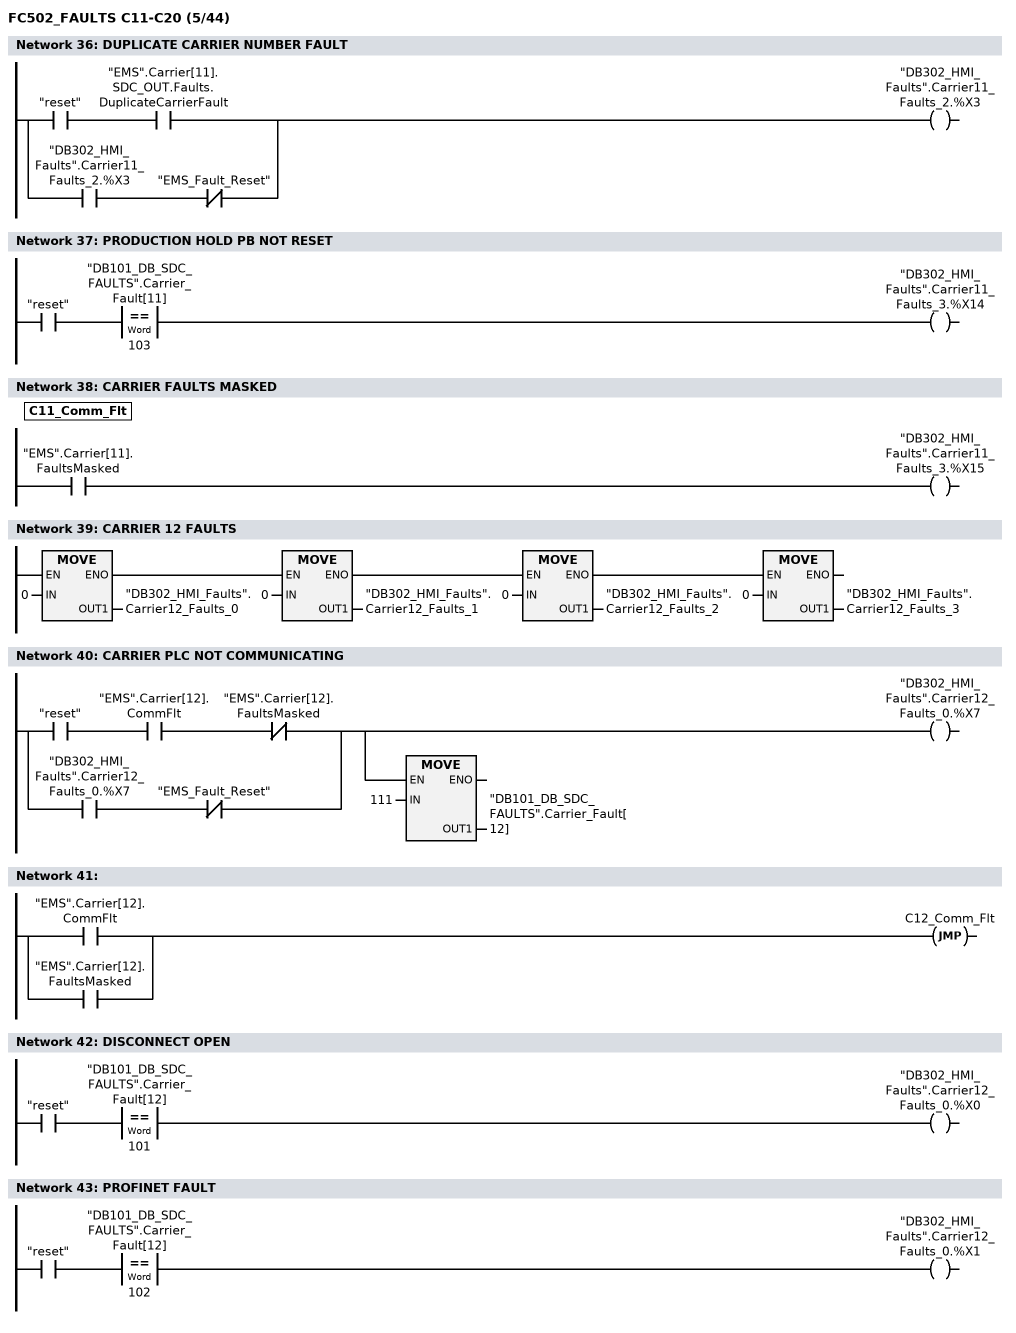
   RUNG wire#powerrail
      Contact( "reset" )
      Contact( "EMS".Carrier[11].SDC_OUT.Faults.DuplicateCarrierFault )
      wire#w1
      Coil( "DB302_HMI_Faults".Carrier11_Faults_2.%X3 )
   END_RUNG
   RUNG wire#powerrail
      Contact( "DB302_HMI_Faults".Carrier11_Faults_2.%X3 )
      I_Contact( "EMS_Fault_Reset" )
   END_RUNG wire#w1
   // the same network as SCL:
   "DB302_HMI_Faults".Carrier11_Faults_2.%X3 := ("reset" AND "EMS".Carrier[11].SDC_OUT.Faults.DuplicateCarrierFault) OR ("DB302_HMI_Faults".Carrier11_Faults_2.%X3 AND NOT "EMS_Fault_Reset");
END_REGION

REGION Network 37: PRODUCTION HOLD PB NOT RESET
   RUNG wire#powerrail
      Contact( "reset" )
      { S7_Templates := "SrcType := Word" } EQ_Contact(in1 := "DB101_DB_SDC_FAULTS".Carrier_Fault[11], in2 := 103)
      Coil( "DB302_HMI_Faults".Carrier11_Faults_3.%X14 )
   END_RUNG
   // the same network as SCL:
   "DB302_HMI_Faults".Carrier11_Faults_3.%X14 := "reset" AND ("DB101_DB_SDC_FAULTS".Carrier_Fault[11] = 103);
END_REGION

REGION Network 38: CARRIER FAULTS MASKED
   Label( C11_Comm_Flt )
   RUNG wire#powerrail
      Contact( "EMS".Carrier[11].FaultsMasked )
      Coil( "DB302_HMI_Faults".Carrier11_Faults_3.%X15 )
   END_RUNG
   // the same network as SCL:
   C11_Comm_Flt:
   "DB302_HMI_Faults".Carrier11_Faults_3.%X15 := "EMS".Carrier[11].FaultsMasked;
END_REGION

REGION Network 39: CARRIER 12 FAULTS
   RUNG wire#powerrail
      Move(in := 0, out1 => "DB302_HMI_Faults".Carrier12_Faults_0)
      Move(in := 0, out1 => "DB302_HMI_Faults".Carrier12_Faults_1)
      Move(in := 0, out1 => "DB302_HMI_Faults".Carrier12_Faults_2)
      Move(in := 0, out1 => "DB302_HMI_Faults".Carrier12_Faults_3)
   END_RUNG
   // the same network as SCL:
   "DB302_HMI_Faults".Carrier12_Faults_0 := 0;
   "DB302_HMI_Faults".Carrier12_Faults_1 := 0;
   "DB302_HMI_Faults".Carrier12_Faults_2 := 0;
   "DB302_HMI_Faults".Carrier12_Faults_3 := 0;
END_REGION

REGION Network 40: CARRIER PLC NOT COMMUNICATING
   RUNG wire#powerrail
      Contact( "reset" )
      Contact( "EMS".Carrier[12].CommFlt )
      I_Contact( "EMS".Carrier[12].FaultsMasked )
      wire#w1
      Coil( "DB302_HMI_Faults".Carrier12_Faults_0.%X7 )
   END_RUNG
   RUNG wire#powerrail
      Contact( "DB302_HMI_Faults".Carrier12_Faults_0.%X7 )
      I_Contact( "EMS_Fault_Reset" )
   END_RUNG wire#w1
   RUNG wire#w1
      Move(in := 111, out1 => "DB101_DB_SDC_FAULTS".Carrier_Fault[12])
   END_RUNG
   // the same network as SCL:
   "DB302_HMI_Faults".Carrier12_Faults_0.%X7 := ("reset" AND "EMS".Carrier[12].CommFlt AND NOT "EMS".Carrier[12].FaultsMasked) OR ("DB302_HMI_Faults".Carrier12_Faults_0.%X7 AND NOT "EMS_Fault_Reset");
   IF "DB302_HMI_Faults".Carrier12_Faults_0.%X7 THEN "DB101_DB_SDC_FAULTS".Carrier_Fault[12] := 111; END_IF;
END_REGION

REGION Network 41
   RUNG wire#powerrail
      Contact( "EMS".Carrier[12].CommFlt )
      wire#w1
      JumpCoil( C12_Comm_Flt )
   END_RUNG
   RUNG wire#powerrail
      Contact( "EMS".Carrier[12].FaultsMasked )
   END_RUNG wire#w1
   // the same network as SCL:
   IF "EMS".Carrier[12].CommFlt OR "EMS".Carrier[12].FaultsMasked THEN GOTO C12_Comm_Flt; END_IF;
END_REGION

REGION Network 42: DISCONNECT OPEN
   RUNG wire#powerrail
      Contact( "reset" )
      { S7_Templates := "SrcType := Word" } EQ_Contact(in1 := "DB101_DB_SDC_FAULTS".Carrier_Fault[12], in2 := 101)
      Coil( "DB302_HMI_Faults".Carrier12_Faults_0.%X0 )
   END_RUNG
   // the same network as SCL:
   "DB302_HMI_Faults".Carrier12_Faults_0.%X0 := "reset" AND ("DB101_DB_SDC_FAULTS".Carrier_Fault[12] = 101);
END_REGION

REGION Network 43: PROFINET FAULT
   RUNG wire#powerrail
      Contact( "reset" )
      { S7_Templates := "SrcType := Word" } EQ_Contact(in1 := "DB101_DB_SDC_FAULTS".Carrier_Fault[12], in2 := 102)
      Coil( "DB302_HMI_Faults".Carrier12_Faults_0.%X1 )
   END_RUNG
   // the same network as SCL:
   "DB302_HMI_Faults".Carrier12_Faults_0.%X1 := "reset" AND ("DB101_DB_SDC_FAULTS".Carrier_Fault[12] = 102);
END_REGION

REGION Network 44: CB2122 TRIPPED
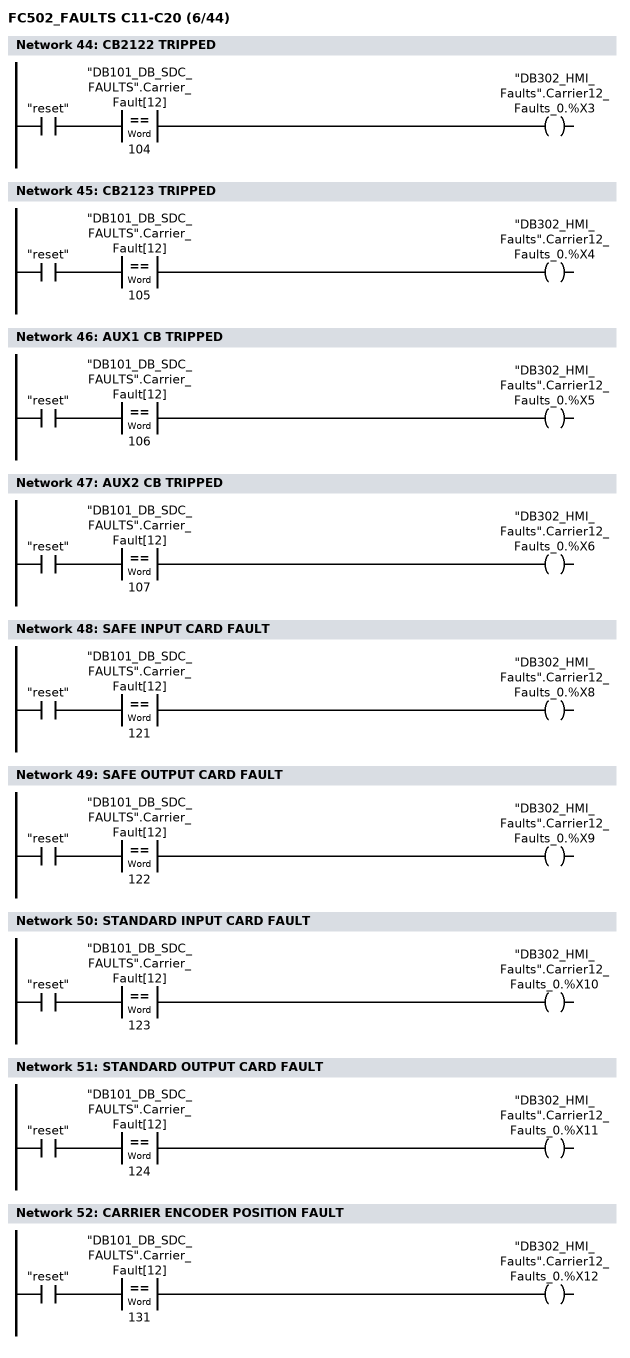
   RUNG wire#powerrail
      Contact( "reset" )
      { S7_Templates := "SrcType := Word" } EQ_Contact(in1 := "DB101_DB_SDC_FAULTS".Carrier_Fault[12], in2 := 104)
      Coil( "DB302_HMI_Faults".Carrier12_Faults_0.%X3 )
   END_RUNG
   // the same network as SCL:
   "DB302_HMI_Faults".Carrier12_Faults_0.%X3 := "reset" AND ("DB101_DB_SDC_FAULTS".Carrier_Fault[12] = 104);
END_REGION

REGION Network 45: CB2123 TRIPPED
   RUNG wire#powerrail
      Contact( "reset" )
      { S7_Templates := "SrcType := Word" } EQ_Contact(in1 := "DB101_DB_SDC_FAULTS".Carrier_Fault[12], in2 := 105)
      Coil( "DB302_HMI_Faults".Carrier12_Faults_0.%X4 )
   END_RUNG
   // the same network as SCL:
   "DB302_HMI_Faults".Carrier12_Faults_0.%X4 := "reset" AND ("DB101_DB_SDC_FAULTS".Carrier_Fault[12] = 105);
END_REGION

REGION Network 46: AUX1 CB TRIPPED
   RUNG wire#powerrail
      Contact( "reset" )
      { S7_Templates := "SrcType := Word" } EQ_Contact(in1 := "DB101_DB_SDC_FAULTS".Carrier_Fault[12], in2 := 106)
      Coil( "DB302_HMI_Faults".Carrier12_Faults_0.%X5 )
   END_RUNG
   // the same network as SCL:
   "DB302_HMI_Faults".Carrier12_Faults_0.%X5 := "reset" AND ("DB101_DB_SDC_FAULTS".Carrier_Fault[12] = 106);
END_REGION

REGION Network 47: AUX2 CB TRIPPED
   RUNG wire#powerrail
      Contact( "reset" )
      { S7_Templates := "SrcType := Word" } EQ_Contact(in1 := "DB101_DB_SDC_FAULTS".Carrier_Fault[12], in2 := 107)
      Coil( "DB302_HMI_Faults".Carrier12_Faults_0.%X6 )
   END_RUNG
   // the same network as SCL:
   "DB302_HMI_Faults".Carrier12_Faults_0.%X6 := "reset" AND ("DB101_DB_SDC_FAULTS".Carrier_Fault[12] = 107);
END_REGION

REGION Network 48: SAFE INPUT CARD FAULT
   RUNG wire#powerrail
      Contact( "reset" )
      { S7_Templates := "SrcType := Word" } EQ_Contact(in1 := "DB101_DB_SDC_FAULTS".Carrier_Fault[12], in2 := 121)
      Coil( "DB302_HMI_Faults".Carrier12_Faults_0.%X8 )
   END_RUNG
   // the same network as SCL:
   "DB302_HMI_Faults".Carrier12_Faults_0.%X8 := "reset" AND ("DB101_DB_SDC_FAULTS".Carrier_Fault[12] = 121);
END_REGION

REGION Network 49: SAFE OUTPUT CARD FAULT
   RUNG wire#powerrail
      Contact( "reset" )
      { S7_Templates := "SrcType := Word" } EQ_Contact(in1 := "DB101_DB_SDC_FAULTS".Carrier_Fault[12], in2 := 122)
      Coil( "DB302_HMI_Faults".Carrier12_Faults_0.%X9 )
   END_RUNG
   // the same network as SCL:
   "DB302_HMI_Faults".Carrier12_Faults_0.%X9 := "reset" AND ("DB101_DB_SDC_FAULTS".Carrier_Fault[12] = 122);
END_REGION

REGION Network 50: STANDARD INPUT CARD FAULT
   RUNG wire#powerrail
      Contact( "reset" )
      { S7_Templates := "SrcType := Word" } EQ_Contact(in1 := "DB101_DB_SDC_FAULTS".Carrier_Fault[12], in2 := 123)
      Coil( "DB302_HMI_Faults".Carrier12_Faults_0.%X10 )
   END_RUNG
   // the same network as SCL:
   "DB302_HMI_Faults".Carrier12_Faults_0.%X10 := "reset" AND ("DB101_DB_SDC_FAULTS".Carrier_Fault[12] = 123);
END_REGION

REGION Network 51: STANDARD OUTPUT CARD FAULT
   RUNG wire#powerrail
      Contact( "reset" )
      { S7_Templates := "SrcType := Word" } EQ_Contact(in1 := "DB101_DB_SDC_FAULTS".Carrier_Fault[12], in2 := 124)
      Coil( "DB302_HMI_Faults".Carrier12_Faults_0.%X11 )
   END_RUNG
   // the same network as SCL:
   "DB302_HMI_Faults".Carrier12_Faults_0.%X11 := "reset" AND ("DB101_DB_SDC_FAULTS".Carrier_Fault[12] = 124);
END_REGION

REGION Network 52: CARRIER ENCODER POSITION FAULT
   RUNG wire#powerrail
      Contact( "reset" )
      { S7_Templates := "SrcType := Word" } EQ_Contact(in1 := "DB101_DB_SDC_FAULTS".Carrier_Fault[12], in2 := 131)
      Coil( "DB302_HMI_Faults".Carrier12_Faults_0.%X12 )
   END_RUNG
   // the same network as SCL:
   "DB302_HMI_Faults".Carrier12_Faults_0.%X12 := "reset" AND ("DB101_DB_SDC_FAULTS".Carrier_Fault[12] = 131);
END_REGION

REGION Network 53: CARRIER ENCODER INTERNAL ERROR
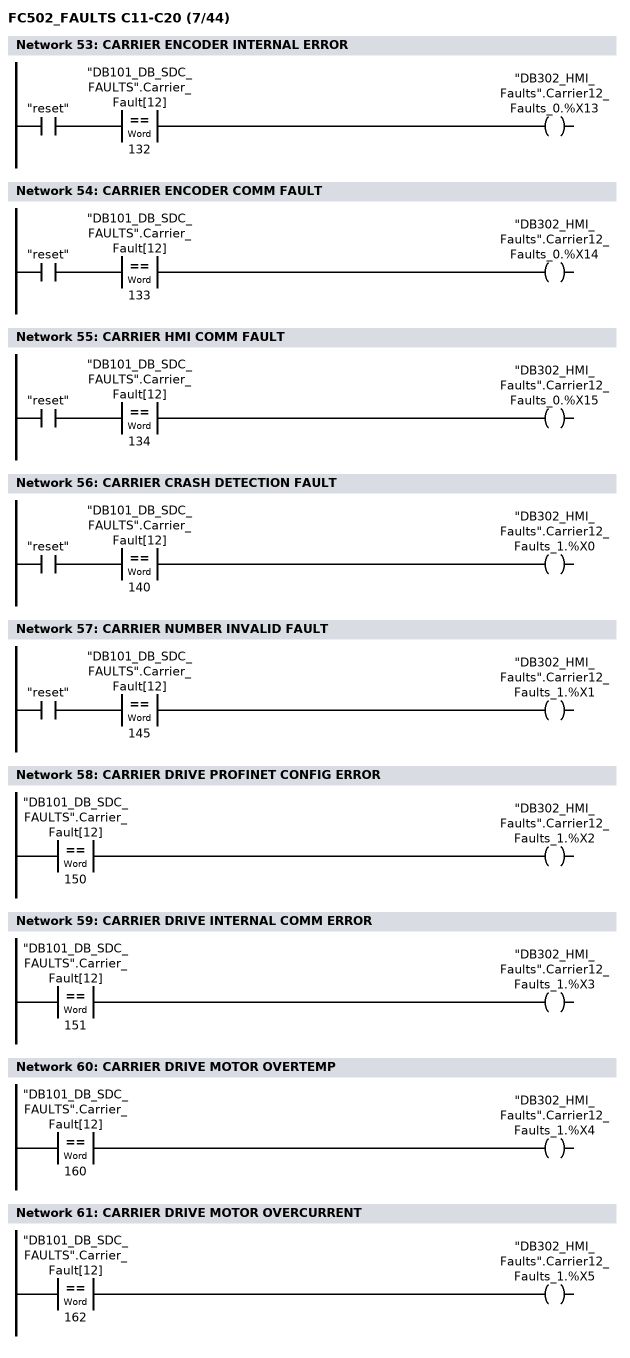
   RUNG wire#powerrail
      Contact( "reset" )
      { S7_Templates := "SrcType := Word" } EQ_Contact(in1 := "DB101_DB_SDC_FAULTS".Carrier_Fault[12], in2 := 132)
      Coil( "DB302_HMI_Faults".Carrier12_Faults_0.%X13 )
   END_RUNG
   // the same network as SCL:
   "DB302_HMI_Faults".Carrier12_Faults_0.%X13 := "reset" AND ("DB101_DB_SDC_FAULTS".Carrier_Fault[12] = 132);
END_REGION

REGION Network 54: CARRIER ENCODER COMM FAULT
   RUNG wire#powerrail
      Contact( "reset" )
      { S7_Templates := "SrcType := Word" } EQ_Contact(in1 := "DB101_DB_SDC_FAULTS".Carrier_Fault[12], in2 := 133)
      Coil( "DB302_HMI_Faults".Carrier12_Faults_0.%X14 )
   END_RUNG
   // the same network as SCL:
   "DB302_HMI_Faults".Carrier12_Faults_0.%X14 := "reset" AND ("DB101_DB_SDC_FAULTS".Carrier_Fault[12] = 133);
END_REGION

REGION Network 55: CARRIER HMI COMM FAULT
   RUNG wire#powerrail
      Contact( "reset" )
      { S7_Templates := "SrcType := Word" } EQ_Contact(in1 := "DB101_DB_SDC_FAULTS".Carrier_Fault[12], in2 := 134)
      Coil( "DB302_HMI_Faults".Carrier12_Faults_0.%X15 )
   END_RUNG
   // the same network as SCL:
   "DB302_HMI_Faults".Carrier12_Faults_0.%X15 := "reset" AND ("DB101_DB_SDC_FAULTS".Carrier_Fault[12] = 134);
END_REGION

REGION Network 56: CARRIER CRASH DETECTION FAULT
   RUNG wire#powerrail
      Contact( "reset" )
      { S7_Templates := "SrcType := Word" } EQ_Contact(in1 := "DB101_DB_SDC_FAULTS".Carrier_Fault[12], in2 := 140)
      Coil( "DB302_HMI_Faults".Carrier12_Faults_1.%X0 )
   END_RUNG
   // the same network as SCL:
   "DB302_HMI_Faults".Carrier12_Faults_1.%X0 := "reset" AND ("DB101_DB_SDC_FAULTS".Carrier_Fault[12] = 140);
END_REGION

REGION Network 57: CARRIER NUMBER INVALID FAULT
   RUNG wire#powerrail
      Contact( "reset" )
      { S7_Templates := "SrcType := Word" } EQ_Contact(in1 := "DB101_DB_SDC_FAULTS".Carrier_Fault[12], in2 := 145)
      Coil( "DB302_HMI_Faults".Carrier12_Faults_1.%X1 )
   END_RUNG
   // the same network as SCL:
   "DB302_HMI_Faults".Carrier12_Faults_1.%X1 := "reset" AND ("DB101_DB_SDC_FAULTS".Carrier_Fault[12] = 145);
END_REGION

REGION Network 58: CARRIER DRIVE PROFINET CONFIG ERROR
   RUNG wire#powerrail
      { S7_Templates := "SrcType := Word" } EQ_Contact(in1 := "DB101_DB_SDC_FAULTS".Carrier_Fault[12], in2 := 150)
      Coil( "DB302_HMI_Faults".Carrier12_Faults_1.%X2 )
   END_RUNG
   // the same network as SCL:
   "DB302_HMI_Faults".Carrier12_Faults_1.%X2 := "DB101_DB_SDC_FAULTS".Carrier_Fault[12] = 150;
END_REGION

REGION Network 59: CARRIER DRIVE INTERNAL COMM ERROR
   RUNG wire#powerrail
      { S7_Templates := "SrcType := Word" } EQ_Contact(in1 := "DB101_DB_SDC_FAULTS".Carrier_Fault[12], in2 := 151)
      Coil( "DB302_HMI_Faults".Carrier12_Faults_1.%X3 )
   END_RUNG
   // the same network as SCL:
   "DB302_HMI_Faults".Carrier12_Faults_1.%X3 := "DB101_DB_SDC_FAULTS".Carrier_Fault[12] = 151;
END_REGION

REGION Network 60: CARRIER DRIVE MOTOR OVERTEMP
   RUNG wire#powerrail
      { S7_Templates := "SrcType := Word" } EQ_Contact(in1 := "DB101_DB_SDC_FAULTS".Carrier_Fault[12], in2 := 160)
      Coil( "DB302_HMI_Faults".Carrier12_Faults_1.%X4 )
   END_RUNG
   // the same network as SCL:
   "DB302_HMI_Faults".Carrier12_Faults_1.%X4 := "DB101_DB_SDC_FAULTS".Carrier_Fault[12] = 160;
END_REGION

REGION Network 61: CARRIER DRIVE MOTOR OVERCURRENT
   RUNG wire#powerrail
      { S7_Templates := "SrcType := Word" } EQ_Contact(in1 := "DB101_DB_SDC_FAULTS".Carrier_Fault[12], in2 := 162)
      Coil( "DB302_HMI_Faults".Carrier12_Faults_1.%X5 )
   END_RUNG
   // the same network as SCL:
   "DB302_HMI_Faults".Carrier12_Faults_1.%X5 := "DB101_DB_SDC_FAULTS".Carrier_Fault[12] = 162;
END_REGION

REGION Network 62: CARRIER DRIVE INFEED OR POWER UNIT NOT READY
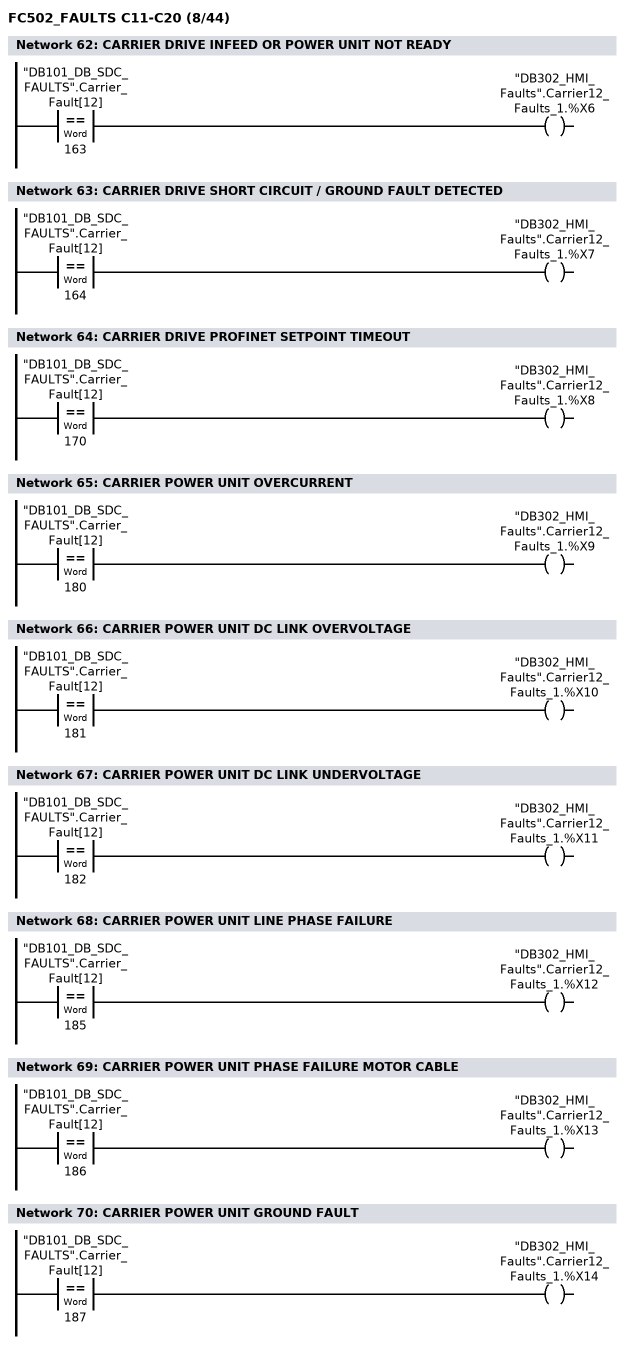
   RUNG wire#powerrail
      { S7_Templates := "SrcType := Word" } EQ_Contact(in1 := "DB101_DB_SDC_FAULTS".Carrier_Fault[12], in2 := 163)
      Coil( "DB302_HMI_Faults".Carrier12_Faults_1.%X6 )
   END_RUNG
   // the same network as SCL:
   "DB302_HMI_Faults".Carrier12_Faults_1.%X6 := "DB101_DB_SDC_FAULTS".Carrier_Fault[12] = 163;
END_REGION

REGION Network 63: CARRIER DRIVE SHORT CIRCUIT / GROUND FAULT DETECTED
   RUNG wire#powerrail
      { S7_Templates := "SrcType := Word" } EQ_Contact(in1 := "DB101_DB_SDC_FAULTS".Carrier_Fault[12], in2 := 164)
      Coil( "DB302_HMI_Faults".Carrier12_Faults_1.%X7 )
   END_RUNG
   // the same network as SCL:
   "DB302_HMI_Faults".Carrier12_Faults_1.%X7 := "DB101_DB_SDC_FAULTS".Carrier_Fault[12] = 164;
END_REGION

REGION Network 64: CARRIER DRIVE PROFINET SETPOINT TIMEOUT
   RUNG wire#powerrail
      { S7_Templates := "SrcType := Word" } EQ_Contact(in1 := "DB101_DB_SDC_FAULTS".Carrier_Fault[12], in2 := 170)
      Coil( "DB302_HMI_Faults".Carrier12_Faults_1.%X8 )
   END_RUNG
   // the same network as SCL:
   "DB302_HMI_Faults".Carrier12_Faults_1.%X8 := "DB101_DB_SDC_FAULTS".Carrier_Fault[12] = 170;
END_REGION

REGION Network 65: CARRIER POWER UNIT OVERCURRENT
   RUNG wire#powerrail
      { S7_Templates := "SrcType := Word" } EQ_Contact(in1 := "DB101_DB_SDC_FAULTS".Carrier_Fault[12], in2 := 180)
      Coil( "DB302_HMI_Faults".Carrier12_Faults_1.%X9 )
   END_RUNG
   // the same network as SCL:
   "DB302_HMI_Faults".Carrier12_Faults_1.%X9 := "DB101_DB_SDC_FAULTS".Carrier_Fault[12] = 180;
END_REGION

REGION Network 66: CARRIER POWER UNIT DC LINK OVERVOLTAGE
   RUNG wire#powerrail
      { S7_Templates := "SrcType := Word" } EQ_Contact(in1 := "DB101_DB_SDC_FAULTS".Carrier_Fault[12], in2 := 181)
      Coil( "DB302_HMI_Faults".Carrier12_Faults_1.%X10 )
   END_RUNG
   // the same network as SCL:
   "DB302_HMI_Faults".Carrier12_Faults_1.%X10 := "DB101_DB_SDC_FAULTS".Carrier_Fault[12] = 181;
END_REGION

REGION Network 67: CARRIER POWER UNIT DC LINK UNDERVOLTAGE
   RUNG wire#powerrail
      { S7_Templates := "SrcType := Word" } EQ_Contact(in1 := "DB101_DB_SDC_FAULTS".Carrier_Fault[12], in2 := 182)
      Coil( "DB302_HMI_Faults".Carrier12_Faults_1.%X11 )
   END_RUNG
   // the same network as SCL:
   "DB302_HMI_Faults".Carrier12_Faults_1.%X11 := "DB101_DB_SDC_FAULTS".Carrier_Fault[12] = 182;
END_REGION

REGION Network 68: CARRIER POWER UNIT LINE PHASE FAILURE
   RUNG wire#powerrail
      { S7_Templates := "SrcType := Word" } EQ_Contact(in1 := "DB101_DB_SDC_FAULTS".Carrier_Fault[12], in2 := 185)
      Coil( "DB302_HMI_Faults".Carrier12_Faults_1.%X12 )
   END_RUNG
   // the same network as SCL:
   "DB302_HMI_Faults".Carrier12_Faults_1.%X12 := "DB101_DB_SDC_FAULTS".Carrier_Fault[12] = 185;
END_REGION

REGION Network 69: CARRIER POWER UNIT PHASE FAILURE MOTOR CABLE
   RUNG wire#powerrail
      { S7_Templates := "SrcType := Word" } EQ_Contact(in1 := "DB101_DB_SDC_FAULTS".Carrier_Fault[12], in2 := 186)
      Coil( "DB302_HMI_Faults".Carrier12_Faults_1.%X13 )
   END_RUNG
   // the same network as SCL:
   "DB302_HMI_Faults".Carrier12_Faults_1.%X13 := "DB101_DB_SDC_FAULTS".Carrier_Fault[12] = 186;
END_REGION

REGION Network 70: CARRIER POWER UNIT GROUND FAULT
   RUNG wire#powerrail
      { S7_Templates := "SrcType := Word" } EQ_Contact(in1 := "DB101_DB_SDC_FAULTS".Carrier_Fault[12], in2 := 187)
      Coil( "DB302_HMI_Faults".Carrier12_Faults_1.%X14 )
   END_RUNG
   // the same network as SCL:
   "DB302_HMI_Faults".Carrier12_Faults_1.%X14 := "DB101_DB_SDC_FAULTS".Carrier_Fault[12] = 187;
END_REGION

REGION Network 71: CARRIER MOTION OFF FAULT
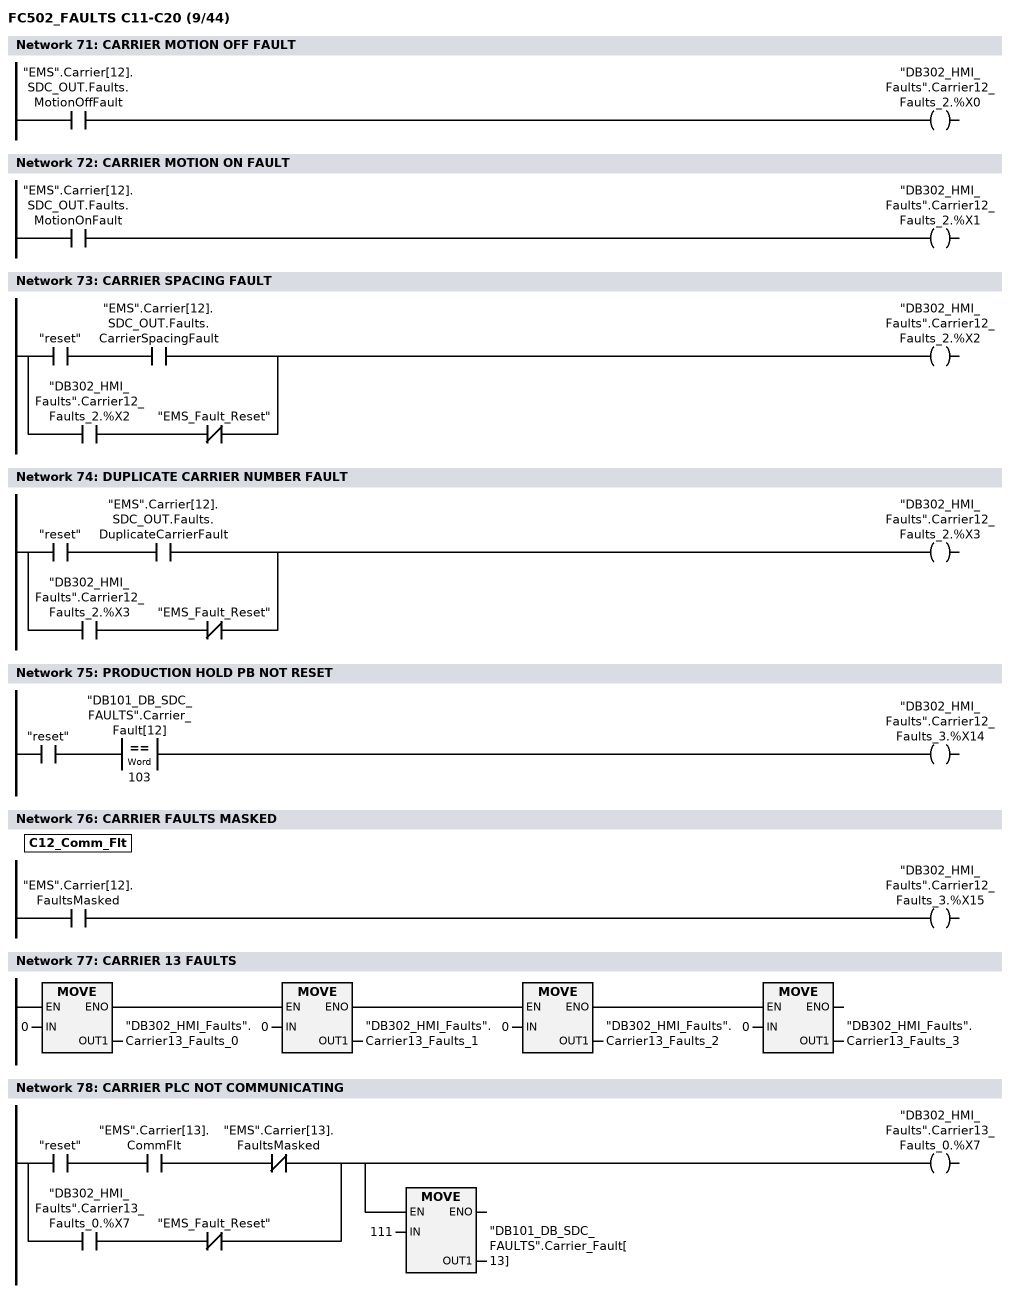
   RUNG wire#powerrail
      Contact( "EMS".Carrier[12].SDC_OUT.Faults.MotionOffFault )
      Coil( "DB302_HMI_Faults".Carrier12_Faults_2.%X0 )
   END_RUNG
   // the same network as SCL:
   "DB302_HMI_Faults".Carrier12_Faults_2.%X0 := "EMS".Carrier[12].SDC_OUT.Faults.MotionOffFault;
END_REGION

REGION Network 72: CARRIER MOTION ON FAULT
   RUNG wire#powerrail
      Contact( "EMS".Carrier[12].SDC_OUT.Faults.MotionOnFault )
      Coil( "DB302_HMI_Faults".Carrier12_Faults_2.%X1 )
   END_RUNG
   // the same network as SCL:
   "DB302_HMI_Faults".Carrier12_Faults_2.%X1 := "EMS".Carrier[12].SDC_OUT.Faults.MotionOnFault;
END_REGION

REGION Network 73: CARRIER SPACING FAULT
   RUNG wire#powerrail
      Contact( "reset" )
      Contact( "EMS".Carrier[12].SDC_OUT.Faults.CarrierSpacingFault )
      wire#w1
      Coil( "DB302_HMI_Faults".Carrier12_Faults_2.%X2 )
   END_RUNG
   RUNG wire#powerrail
      Contact( "DB302_HMI_Faults".Carrier12_Faults_2.%X2 )
      I_Contact( "EMS_Fault_Reset" )
   END_RUNG wire#w1
   // the same network as SCL:
   "DB302_HMI_Faults".Carrier12_Faults_2.%X2 := ("reset" AND "EMS".Carrier[12].SDC_OUT.Faults.CarrierSpacingFault) OR ("DB302_HMI_Faults".Carrier12_Faults_2.%X2 AND NOT "EMS_Fault_Reset");
END_REGION

REGION Network 74: DUPLICATE CARRIER NUMBER FAULT
   RUNG wire#powerrail
      Contact( "reset" )
      Contact( "EMS".Carrier[12].SDC_OUT.Faults.DuplicateCarrierFault )
      wire#w1
      Coil( "DB302_HMI_Faults".Carrier12_Faults_2.%X3 )
   END_RUNG
   RUNG wire#powerrail
      Contact( "DB302_HMI_Faults".Carrier12_Faults_2.%X3 )
      I_Contact( "EMS_Fault_Reset" )
   END_RUNG wire#w1
   // the same network as SCL:
   "DB302_HMI_Faults".Carrier12_Faults_2.%X3 := ("reset" AND "EMS".Carrier[12].SDC_OUT.Faults.DuplicateCarrierFault) OR ("DB302_HMI_Faults".Carrier12_Faults_2.%X3 AND NOT "EMS_Fault_Reset");
END_REGION

REGION Network 75: PRODUCTION HOLD PB NOT RESET
   RUNG wire#powerrail
      Contact( "reset" )
      { S7_Templates := "SrcType := Word" } EQ_Contact(in1 := "DB101_DB_SDC_FAULTS".Carrier_Fault[12], in2 := 103)
      Coil( "DB302_HMI_Faults".Carrier12_Faults_3.%X14 )
   END_RUNG
   // the same network as SCL:
   "DB302_HMI_Faults".Carrier12_Faults_3.%X14 := "reset" AND ("DB101_DB_SDC_FAULTS".Carrier_Fault[12] = 103);
END_REGION

REGION Network 76: CARRIER FAULTS MASKED
   Label( C12_Comm_Flt )
   RUNG wire#powerrail
      Contact( "EMS".Carrier[12].FaultsMasked )
      Coil( "DB302_HMI_Faults".Carrier12_Faults_3.%X15 )
   END_RUNG
   // the same network as SCL:
   C12_Comm_Flt:
   "DB302_HMI_Faults".Carrier12_Faults_3.%X15 := "EMS".Carrier[12].FaultsMasked;
END_REGION

REGION Network 77: CARRIER 13 FAULTS
   RUNG wire#powerrail
      Move(in := 0, out1 => "DB302_HMI_Faults".Carrier13_Faults_0)
      Move(in := 0, out1 => "DB302_HMI_Faults".Carrier13_Faults_1)
      Move(in := 0, out1 => "DB302_HMI_Faults".Carrier13_Faults_2)
      Move(in := 0, out1 => "DB302_HMI_Faults".Carrier13_Faults_3)
   END_RUNG
   // the same network as SCL:
   "DB302_HMI_Faults".Carrier13_Faults_0 := 0;
   "DB302_HMI_Faults".Carrier13_Faults_1 := 0;
   "DB302_HMI_Faults".Carrier13_Faults_2 := 0;
   "DB302_HMI_Faults".Carrier13_Faults_3 := 0;
END_REGION

REGION Network 78: CARRIER PLC NOT COMMUNICATING
   RUNG wire#powerrail
      Contact( "reset" )
      Contact( "EMS".Carrier[13].CommFlt )
      I_Contact( "EMS".Carrier[13].FaultsMasked )
      wire#w1
      Coil( "DB302_HMI_Faults".Carrier13_Faults_0.%X7 )
   END_RUNG
   RUNG wire#powerrail
      Contact( "DB302_HMI_Faults".Carrier13_Faults_0.%X7 )
      I_Contact( "EMS_Fault_Reset" )
   END_RUNG wire#w1
   RUNG wire#w1
      Move(in := 111, out1 => "DB101_DB_SDC_FAULTS".Carrier_Fault[13])
   END_RUNG
   // the same network as SCL:
   "DB302_HMI_Faults".Carrier13_Faults_0.%X7 := ("reset" AND "EMS".Carrier[13].CommFlt AND NOT "EMS".Carrier[13].FaultsMasked) OR ("DB302_HMI_Faults".Carrier13_Faults_0.%X7 AND NOT "EMS_Fault_Reset");
   IF "DB302_HMI_Faults".Carrier13_Faults_0.%X7 THEN "DB101_DB_SDC_FAULTS".Carrier_Fault[13] := 111; END_IF;
END_REGION

REGION Network 79
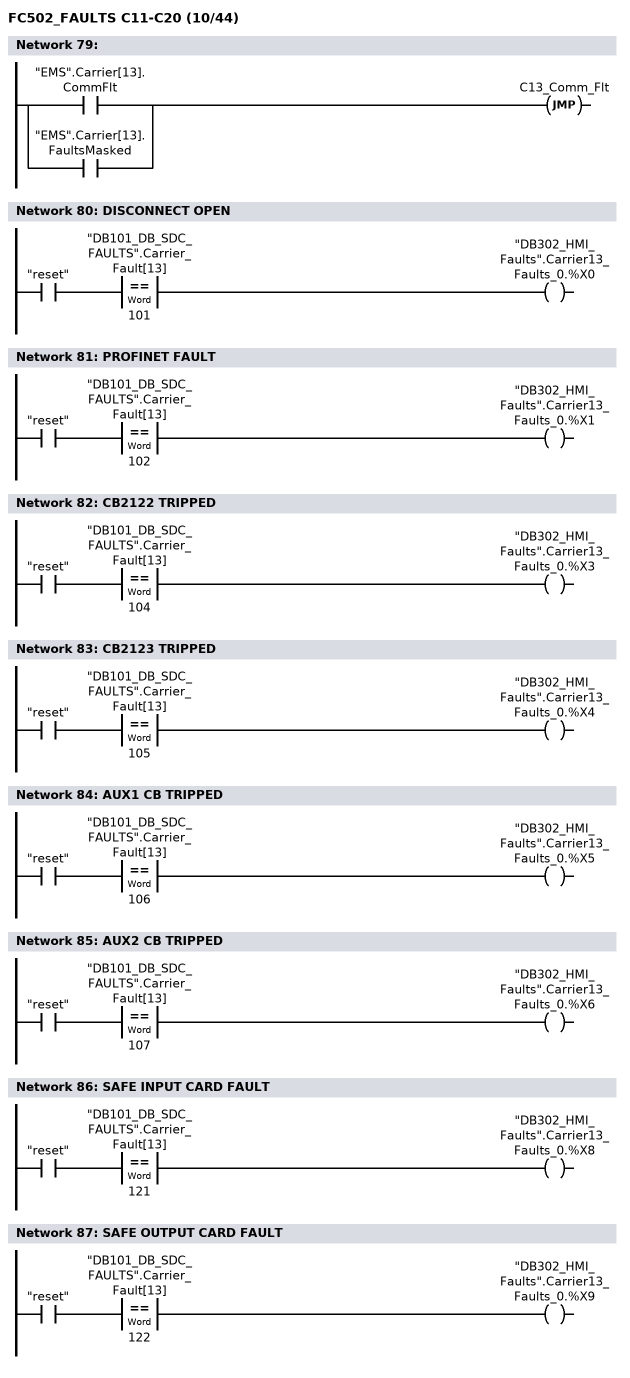
   RUNG wire#powerrail
      Contact( "EMS".Carrier[13].CommFlt )
      wire#w1
      JumpCoil( C13_Comm_Flt )
   END_RUNG
   RUNG wire#powerrail
      Contact( "EMS".Carrier[13].FaultsMasked )
   END_RUNG wire#w1
   // the same network as SCL:
   IF "EMS".Carrier[13].CommFlt OR "EMS".Carrier[13].FaultsMasked THEN GOTO C13_Comm_Flt; END_IF;
END_REGION

REGION Network 80: DISCONNECT OPEN
   RUNG wire#powerrail
      Contact( "reset" )
      { S7_Templates := "SrcType := Word" } EQ_Contact(in1 := "DB101_DB_SDC_FAULTS".Carrier_Fault[13], in2 := 101)
      Coil( "DB302_HMI_Faults".Carrier13_Faults_0.%X0 )
   END_RUNG
   // the same network as SCL:
   "DB302_HMI_Faults".Carrier13_Faults_0.%X0 := "reset" AND ("DB101_DB_SDC_FAULTS".Carrier_Fault[13] = 101);
END_REGION

REGION Network 81: PROFINET FAULT
   RUNG wire#powerrail
      Contact( "reset" )
      { S7_Templates := "SrcType := Word" } EQ_Contact(in1 := "DB101_DB_SDC_FAULTS".Carrier_Fault[13], in2 := 102)
      Coil( "DB302_HMI_Faults".Carrier13_Faults_0.%X1 )
   END_RUNG
   // the same network as SCL:
   "DB302_HMI_Faults".Carrier13_Faults_0.%X1 := "reset" AND ("DB101_DB_SDC_FAULTS".Carrier_Fault[13] = 102);
END_REGION

REGION Network 82: CB2122 TRIPPED
   RUNG wire#powerrail
      Contact( "reset" )
      { S7_Templates := "SrcType := Word" } EQ_Contact(in1 := "DB101_DB_SDC_FAULTS".Carrier_Fault[13], in2 := 104)
      Coil( "DB302_HMI_Faults".Carrier13_Faults_0.%X3 )
   END_RUNG
   // the same network as SCL:
   "DB302_HMI_Faults".Carrier13_Faults_0.%X3 := "reset" AND ("DB101_DB_SDC_FAULTS".Carrier_Fault[13] = 104);
END_REGION

REGION Network 83: CB2123 TRIPPED
   RUNG wire#powerrail
      Contact( "reset" )
      { S7_Templates := "SrcType := Word" } EQ_Contact(in1 := "DB101_DB_SDC_FAULTS".Carrier_Fault[13], in2 := 105)
      Coil( "DB302_HMI_Faults".Carrier13_Faults_0.%X4 )
   END_RUNG
   // the same network as SCL:
   "DB302_HMI_Faults".Carrier13_Faults_0.%X4 := "reset" AND ("DB101_DB_SDC_FAULTS".Carrier_Fault[13] = 105);
END_REGION

REGION Network 84: AUX1 CB TRIPPED
   RUNG wire#powerrail
      Contact( "reset" )
      { S7_Templates := "SrcType := Word" } EQ_Contact(in1 := "DB101_DB_SDC_FAULTS".Carrier_Fault[13], in2 := 106)
      Coil( "DB302_HMI_Faults".Carrier13_Faults_0.%X5 )
   END_RUNG
   // the same network as SCL:
   "DB302_HMI_Faults".Carrier13_Faults_0.%X5 := "reset" AND ("DB101_DB_SDC_FAULTS".Carrier_Fault[13] = 106);
END_REGION

REGION Network 85: AUX2 CB TRIPPED
   RUNG wire#powerrail
      Contact( "reset" )
      { S7_Templates := "SrcType := Word" } EQ_Contact(in1 := "DB101_DB_SDC_FAULTS".Carrier_Fault[13], in2 := 107)
      Coil( "DB302_HMI_Faults".Carrier13_Faults_0.%X6 )
   END_RUNG
   // the same network as SCL:
   "DB302_HMI_Faults".Carrier13_Faults_0.%X6 := "reset" AND ("DB101_DB_SDC_FAULTS".Carrier_Fault[13] = 107);
END_REGION

REGION Network 86: SAFE INPUT CARD FAULT
   RUNG wire#powerrail
      Contact( "reset" )
      { S7_Templates := "SrcType := Word" } EQ_Contact(in1 := "DB101_DB_SDC_FAULTS".Carrier_Fault[13], in2 := 121)
      Coil( "DB302_HMI_Faults".Carrier13_Faults_0.%X8 )
   END_RUNG
   // the same network as SCL:
   "DB302_HMI_Faults".Carrier13_Faults_0.%X8 := "reset" AND ("DB101_DB_SDC_FAULTS".Carrier_Fault[13] = 121);
END_REGION

REGION Network 87: SAFE OUTPUT CARD FAULT
   RUNG wire#powerrail
      Contact( "reset" )
      { S7_Templates := "SrcType := Word" } EQ_Contact(in1 := "DB101_DB_SDC_FAULTS".Carrier_Fault[13], in2 := 122)
      Coil( "DB302_HMI_Faults".Carrier13_Faults_0.%X9 )
   END_RUNG
   // the same network as SCL:
   "DB302_HMI_Faults".Carrier13_Faults_0.%X9 := "reset" AND ("DB101_DB_SDC_FAULTS".Carrier_Fault[13] = 122);
END_REGION

REGION Network 88: STANDARD INPUT CARD FAULT
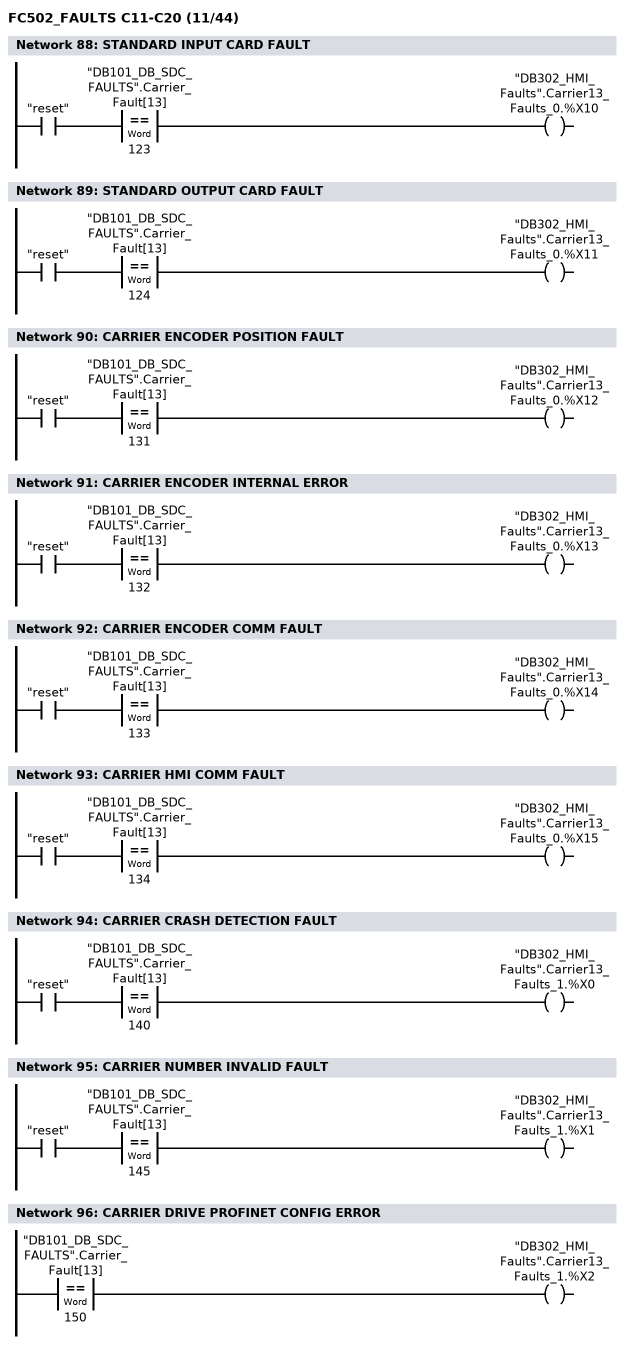
   RUNG wire#powerrail
      Contact( "reset" )
      { S7_Templates := "SrcType := Word" } EQ_Contact(in1 := "DB101_DB_SDC_FAULTS".Carrier_Fault[13], in2 := 123)
      Coil( "DB302_HMI_Faults".Carrier13_Faults_0.%X10 )
   END_RUNG
   // the same network as SCL:
   "DB302_HMI_Faults".Carrier13_Faults_0.%X10 := "reset" AND ("DB101_DB_SDC_FAULTS".Carrier_Fault[13] = 123);
END_REGION

REGION Network 89: STANDARD OUTPUT CARD FAULT
   RUNG wire#powerrail
      Contact( "reset" )
      { S7_Templates := "SrcType := Word" } EQ_Contact(in1 := "DB101_DB_SDC_FAULTS".Carrier_Fault[13], in2 := 124)
      Coil( "DB302_HMI_Faults".Carrier13_Faults_0.%X11 )
   END_RUNG
   // the same network as SCL:
   "DB302_HMI_Faults".Carrier13_Faults_0.%X11 := "reset" AND ("DB101_DB_SDC_FAULTS".Carrier_Fault[13] = 124);
END_REGION

REGION Network 90: CARRIER ENCODER POSITION FAULT
   RUNG wire#powerrail
      Contact( "reset" )
      { S7_Templates := "SrcType := Word" } EQ_Contact(in1 := "DB101_DB_SDC_FAULTS".Carrier_Fault[13], in2 := 131)
      Coil( "DB302_HMI_Faults".Carrier13_Faults_0.%X12 )
   END_RUNG
   // the same network as SCL:
   "DB302_HMI_Faults".Carrier13_Faults_0.%X12 := "reset" AND ("DB101_DB_SDC_FAULTS".Carrier_Fault[13] = 131);
END_REGION

REGION Network 91: CARRIER ENCODER INTERNAL ERROR
   RUNG wire#powerrail
      Contact( "reset" )
      { S7_Templates := "SrcType := Word" } EQ_Contact(in1 := "DB101_DB_SDC_FAULTS".Carrier_Fault[13], in2 := 132)
      Coil( "DB302_HMI_Faults".Carrier13_Faults_0.%X13 )
   END_RUNG
   // the same network as SCL:
   "DB302_HMI_Faults".Carrier13_Faults_0.%X13 := "reset" AND ("DB101_DB_SDC_FAULTS".Carrier_Fault[13] = 132);
END_REGION

REGION Network 92: CARRIER ENCODER COMM FAULT
   RUNG wire#powerrail
      Contact( "reset" )
      { S7_Templates := "SrcType := Word" } EQ_Contact(in1 := "DB101_DB_SDC_FAULTS".Carrier_Fault[13], in2 := 133)
      Coil( "DB302_HMI_Faults".Carrier13_Faults_0.%X14 )
   END_RUNG
   // the same network as SCL:
   "DB302_HMI_Faults".Carrier13_Faults_0.%X14 := "reset" AND ("DB101_DB_SDC_FAULTS".Carrier_Fault[13] = 133);
END_REGION

REGION Network 93: CARRIER HMI COMM FAULT
   RUNG wire#powerrail
      Contact( "reset" )
      { S7_Templates := "SrcType := Word" } EQ_Contact(in1 := "DB101_DB_SDC_FAULTS".Carrier_Fault[13], in2 := 134)
      Coil( "DB302_HMI_Faults".Carrier13_Faults_0.%X15 )
   END_RUNG
   // the same network as SCL:
   "DB302_HMI_Faults".Carrier13_Faults_0.%X15 := "reset" AND ("DB101_DB_SDC_FAULTS".Carrier_Fault[13] = 134);
END_REGION

REGION Network 94: CARRIER CRASH DETECTION FAULT
   RUNG wire#powerrail
      Contact( "reset" )
      { S7_Templates := "SrcType := Word" } EQ_Contact(in1 := "DB101_DB_SDC_FAULTS".Carrier_Fault[13], in2 := 140)
      Coil( "DB302_HMI_Faults".Carrier13_Faults_1.%X0 )
   END_RUNG
   // the same network as SCL:
   "DB302_HMI_Faults".Carrier13_Faults_1.%X0 := "reset" AND ("DB101_DB_SDC_FAULTS".Carrier_Fault[13] = 140);
END_REGION

REGION Network 95: CARRIER NUMBER INVALID FAULT
   RUNG wire#powerrail
      Contact( "reset" )
      { S7_Templates := "SrcType := Word" } EQ_Contact(in1 := "DB101_DB_SDC_FAULTS".Carrier_Fault[13], in2 := 145)
      Coil( "DB302_HMI_Faults".Carrier13_Faults_1.%X1 )
   END_RUNG
   // the same network as SCL:
   "DB302_HMI_Faults".Carrier13_Faults_1.%X1 := "reset" AND ("DB101_DB_SDC_FAULTS".Carrier_Fault[13] = 145);
END_REGION

REGION Network 96: CARRIER DRIVE PROFINET CONFIG ERROR
   RUNG wire#powerrail
      { S7_Templates := "SrcType := Word" } EQ_Contact(in1 := "DB101_DB_SDC_FAULTS".Carrier_Fault[13], in2 := 150)
      Coil( "DB302_HMI_Faults".Carrier13_Faults_1.%X2 )
   END_RUNG
   // the same network as SCL:
   "DB302_HMI_Faults".Carrier13_Faults_1.%X2 := "DB101_DB_SDC_FAULTS".Carrier_Fault[13] = 150;
END_REGION

REGION Network 97: CARRIER DRIVE INTERNAL COMM ERROR
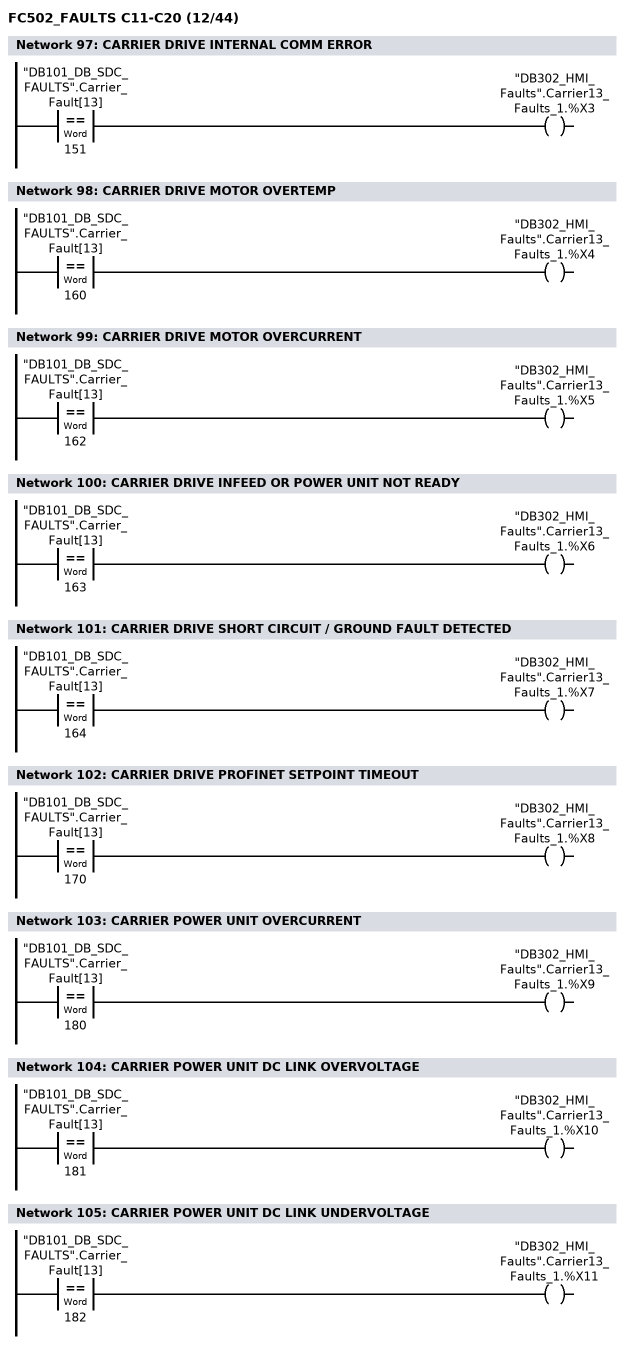
   RUNG wire#powerrail
      { S7_Templates := "SrcType := Word" } EQ_Contact(in1 := "DB101_DB_SDC_FAULTS".Carrier_Fault[13], in2 := 151)
      Coil( "DB302_HMI_Faults".Carrier13_Faults_1.%X3 )
   END_RUNG
   // the same network as SCL:
   "DB302_HMI_Faults".Carrier13_Faults_1.%X3 := "DB101_DB_SDC_FAULTS".Carrier_Fault[13] = 151;
END_REGION

REGION Network 98: CARRIER DRIVE MOTOR OVERTEMP
   RUNG wire#powerrail
      { S7_Templates := "SrcType := Word" } EQ_Contact(in1 := "DB101_DB_SDC_FAULTS".Carrier_Fault[13], in2 := 160)
      Coil( "DB302_HMI_Faults".Carrier13_Faults_1.%X4 )
   END_RUNG
   // the same network as SCL:
   "DB302_HMI_Faults".Carrier13_Faults_1.%X4 := "DB101_DB_SDC_FAULTS".Carrier_Fault[13] = 160;
END_REGION

REGION Network 99: CARRIER DRIVE MOTOR OVERCURRENT
   RUNG wire#powerrail
      { S7_Templates := "SrcType := Word" } EQ_Contact(in1 := "DB101_DB_SDC_FAULTS".Carrier_Fault[13], in2 := 162)
      Coil( "DB302_HMI_Faults".Carrier13_Faults_1.%X5 )
   END_RUNG
   // the same network as SCL:
   "DB302_HMI_Faults".Carrier13_Faults_1.%X5 := "DB101_DB_SDC_FAULTS".Carrier_Fault[13] = 162;
END_REGION

REGION Network 100: CARRIER DRIVE INFEED OR POWER UNIT NOT READY
   RUNG wire#powerrail
      { S7_Templates := "SrcType := Word" } EQ_Contact(in1 := "DB101_DB_SDC_FAULTS".Carrier_Fault[13], in2 := 163)
      Coil( "DB302_HMI_Faults".Carrier13_Faults_1.%X6 )
   END_RUNG
   // the same network as SCL:
   "DB302_HMI_Faults".Carrier13_Faults_1.%X6 := "DB101_DB_SDC_FAULTS".Carrier_Fault[13] = 163;
END_REGION

REGION Network 101: CARRIER DRIVE SHORT CIRCUIT / GROUND FAULT DETECTED
   RUNG wire#powerrail
      { S7_Templates := "SrcType := Word" } EQ_Contact(in1 := "DB101_DB_SDC_FAULTS".Carrier_Fault[13], in2 := 164)
      Coil( "DB302_HMI_Faults".Carrier13_Faults_1.%X7 )
   END_RUNG
   // the same network as SCL:
   "DB302_HMI_Faults".Carrier13_Faults_1.%X7 := "DB101_DB_SDC_FAULTS".Carrier_Fault[13] = 164;
END_REGION

REGION Network 102: CARRIER DRIVE PROFINET SETPOINT TIMEOUT
   RUNG wire#powerrail
      { S7_Templates := "SrcType := Word" } EQ_Contact(in1 := "DB101_DB_SDC_FAULTS".Carrier_Fault[13], in2 := 170)
      Coil( "DB302_HMI_Faults".Carrier13_Faults_1.%X8 )
   END_RUNG
   // the same network as SCL:
   "DB302_HMI_Faults".Carrier13_Faults_1.%X8 := "DB101_DB_SDC_FAULTS".Carrier_Fault[13] = 170;
END_REGION

REGION Network 103: CARRIER POWER UNIT OVERCURRENT
   RUNG wire#powerrail
      { S7_Templates := "SrcType := Word" } EQ_Contact(in1 := "DB101_DB_SDC_FAULTS".Carrier_Fault[13], in2 := 180)
      Coil( "DB302_HMI_Faults".Carrier13_Faults_1.%X9 )
   END_RUNG
   // the same network as SCL:
   "DB302_HMI_Faults".Carrier13_Faults_1.%X9 := "DB101_DB_SDC_FAULTS".Carrier_Fault[13] = 180;
END_REGION

REGION Network 104: CARRIER POWER UNIT DC LINK OVERVOLTAGE
   RUNG wire#powerrail
      { S7_Templates := "SrcType := Word" } EQ_Contact(in1 := "DB101_DB_SDC_FAULTS".Carrier_Fault[13], in2 := 181)
      Coil( "DB302_HMI_Faults".Carrier13_Faults_1.%X10 )
   END_RUNG
   // the same network as SCL:
   "DB302_HMI_Faults".Carrier13_Faults_1.%X10 := "DB101_DB_SDC_FAULTS".Carrier_Fault[13] = 181;
END_REGION

REGION Network 105: CARRIER POWER UNIT DC LINK UNDERVOLTAGE
   RUNG wire#powerrail
      { S7_Templates := "SrcType := Word" } EQ_Contact(in1 := "DB101_DB_SDC_FAULTS".Carrier_Fault[13], in2 := 182)
      Coil( "DB302_HMI_Faults".Carrier13_Faults_1.%X11 )
   END_RUNG
   // the same network as SCL:
   "DB302_HMI_Faults".Carrier13_Faults_1.%X11 := "DB101_DB_SDC_FAULTS".Carrier_Fault[13] = 182;
END_REGION

REGION Network 106: CARRIER POWER UNIT LINE PHASE FAILURE